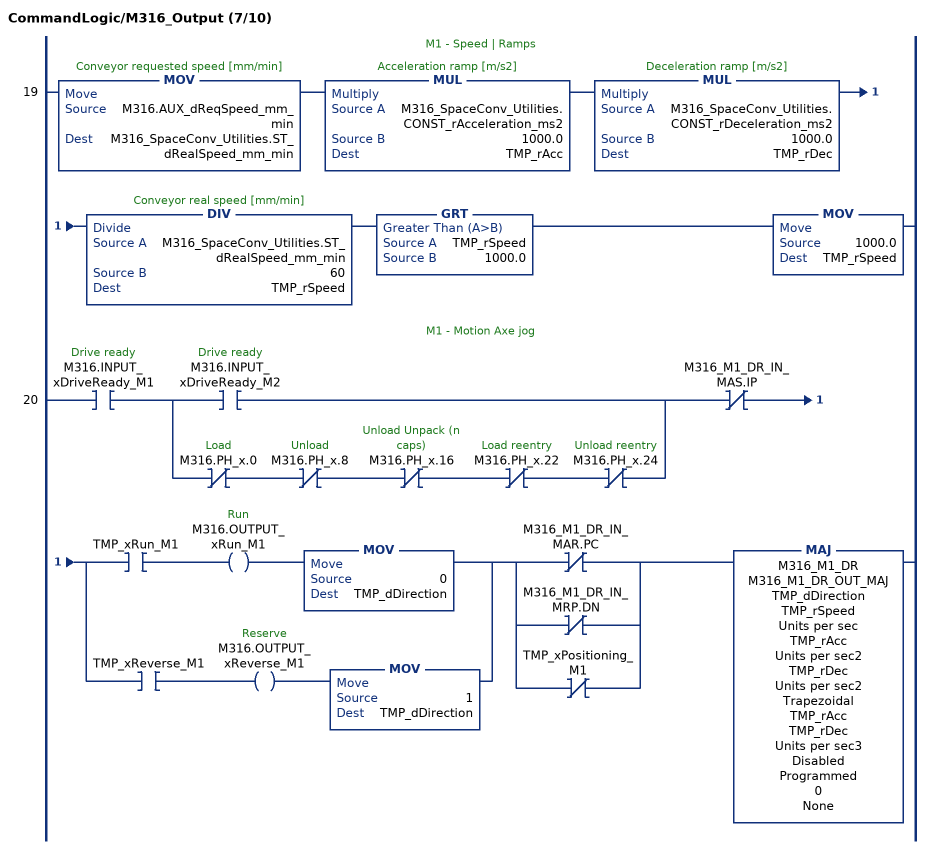
   // M1 - Speed | Ramps
   19: MOV(M316.AUX_dReqSpeed_mm_min,M316_SpaceConv_Utilities.ST_dRealSpeed_mm_min)MUL(M316_SpaceConv_Utilities.CONST_rAcceleration_ms2,1000.0,TMP_rAcc)MUL(M316_SpaceConv_Utilities.CONST_rDeceleration_ms2,1000.0,TMP_rDec)DIV(M316_SpaceConv_Utilities.ST_dRealSpeed_mm_min,60,TMP_rSpeed)GRT(TMP_rSpeed,1000.0)MOV(1000.0,TMP_rSpeed);
   // M1 - Motion Axe jog
   20: XIC(M316.INPUT_xDriveReady_M1)[XIC(M316.INPUT_xDriveReady_M2) ,XIO(M316.PH_x.0) XIO(M316.PH_x.8) XIO(M316.PH_x.16) XIO(M316.PH_x.22) XIO(M316.PH_x.24) ]XIO(M316_M1_DR_IN_MAS.IP)[XIC(TMP_xRun_M1) OTE(M316.OUTPUT_xRun_M1) MOV(0,TMP_dDirection) ,XIC(TMP_xReverse_M1) OTE(M316.OUTPUT_xReverse_M1) MOV(1,TMP_dDirection) ][XIO(M316_M1_DR_IN_MAR.PC) ,XIO(M316_M1_DR_IN_MRP.DN) ,XIO(TMP_xPositioning_M1) ]MAJ(M316_M1_DR,M316_M1_DR_OUT_MAJ,TMP_dDirection,TMP_rSpeed,Units per sec,TMP_rAcc,Units per sec2,TMP_rDec,Units per sec2,Trapezoidal,TMP_rAcc,TMP_rDec,Units per sec3,Disabled,Programmed,0,None);
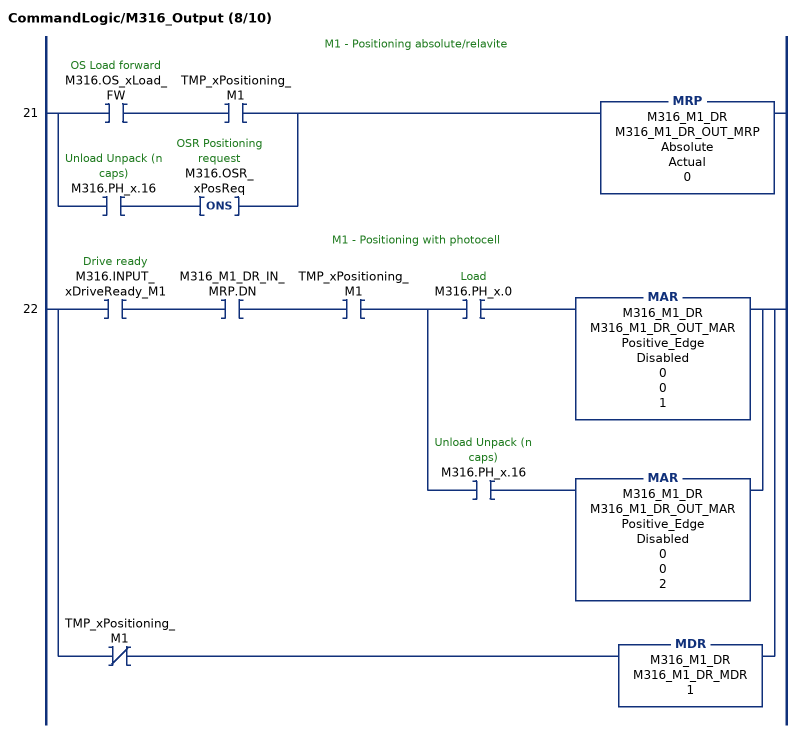
   // M1 - Positioning absolute/relavite
   21: [XIC(M316.OS_xLoad_FW) XIC(TMP_xPositioning_M1) ,XIC(M316.PH_x.16) ONS(M316.OSR_xPosReq) ]MRP(M316_M1_DR,M316_M1_DR_OUT_MRP,Absolute,Actual,0);
   // M1 - Positioning with photocell
   22: [XIC(M316.INPUT_xDriveReady_M1) XIC(M316_M1_DR_IN_MRP.DN) XIC(TMP_xPositioning_M1) [XIC(M316.PH_x.0) MAR(M316_M1_DR,M316_M1_DR_OUT_MAR,Positive_Edge,Disabled,0,0,1) ,XIC(M316.PH_x.16) MAR(M316_M1_DR,M316_M1_DR_OUT_MAR,Positive_Edge,Disabled,0,0,2) ] ,XIO(TMP_xPositioning_M1) MDR(M316_M1_DR,M316_M1_DR_MDR,1) ];
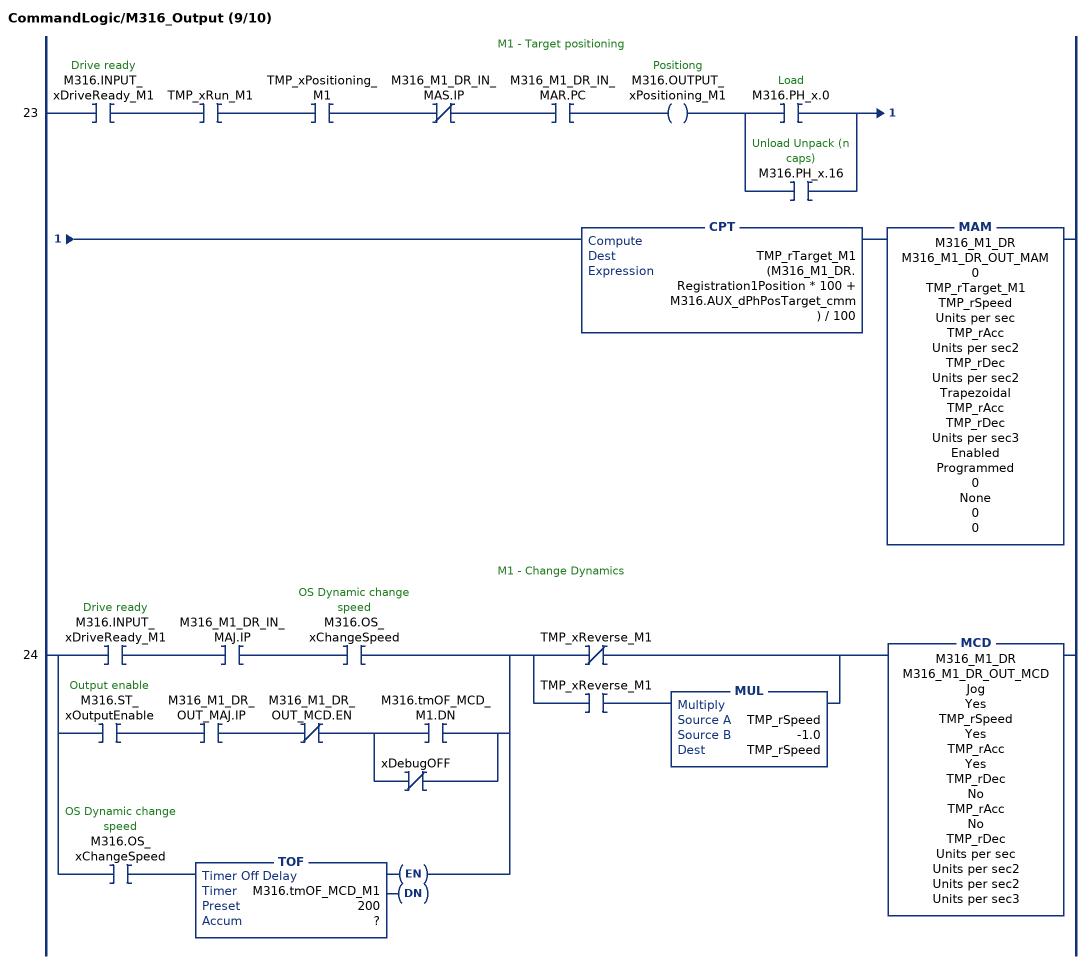
   // M1 - Target positioning
   23: XIC(M316.INPUT_xDriveReady_M1)XIC(TMP_xRun_M1)XIC(TMP_xPositioning_M1)XIO(M316_M1_DR_IN_MAS.IP)XIC(M316_M1_DR_IN_MAR.PC)OTE(M316.OUTPUT_xPositioning_M1)[XIC(M316.PH_x.0) ,XIC(M316.PH_x.16) ]CPT(TMP_rTarget_M1,(M316_M1_DR.Registration1Position * 100 + M316.AUX_dPhPosTarget_cmm ) / 100)MAM(M316_M1_DR,M316_M1_DR_OUT_MAM,0,TMP_rTarget_M1,TMP_rSpeed,Units per sec,TMP_rAcc,Units per sec2,TMP_rDec,Units per sec2,Trapezoidal,TMP_rAcc,TMP_rDec,Units per sec3,Enabled,Programmed,0,None,0,0);
   // M1 - Change Dynamics
   24: [XIC(M316.INPUT_xDriveReady_M1) XIC(M316_M1_DR_IN_MAJ.IP) XIC(M316.OS_xChangeSpeed) ,XIC(M316.ST_xOutputEnable) XIC(M316_M1_DR_OUT_MAJ.IP) XIO(M316_M1_DR_OUT_MCD.EN) [XIC(M316.tmOF_MCD_M1.DN) ,XIO(xDebugOFF) ] ,XIC(M316.OS_xChangeSpeed) TOF(M316.tmOF_MCD_M1,?,?) ][XIO(TMP_xReverse_M1) ,XIC(TMP_xReverse_M1) MUL(TMP_rSpeed,-1.0,TMP_rSpeed) ]MCD(M316_M1_DR,M316_M1_DR_OUT_MCD,Jog,Yes,TMP_rSpeed,Yes,TMP_rAcc,Yes,TMP_rDec,No,TMP_rAcc,No,TMP_rDec,Units per sec,Units per sec2,Units per sec2,Units per sec3);
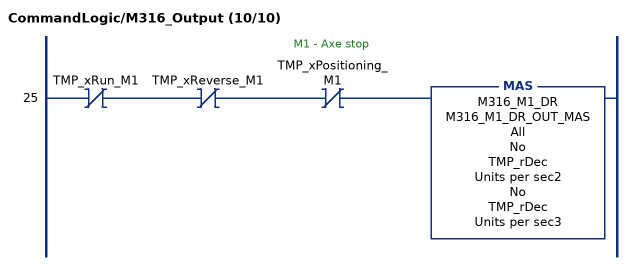
   // M1 - Axe stop
   25: XIO(TMP_xRun_M1)XIO(TMP_xReverse_M1)XIO(TMP_xPositioning_M1)MAS(M316_M1_DR,M316_M1_DR_OUT_MAS,All,No,TMP_rDec,Units per sec2,No,TMP_rDec,Units per sec3);
END_ROUTINE

ROUTINE M316A_Output   (* ladder *)
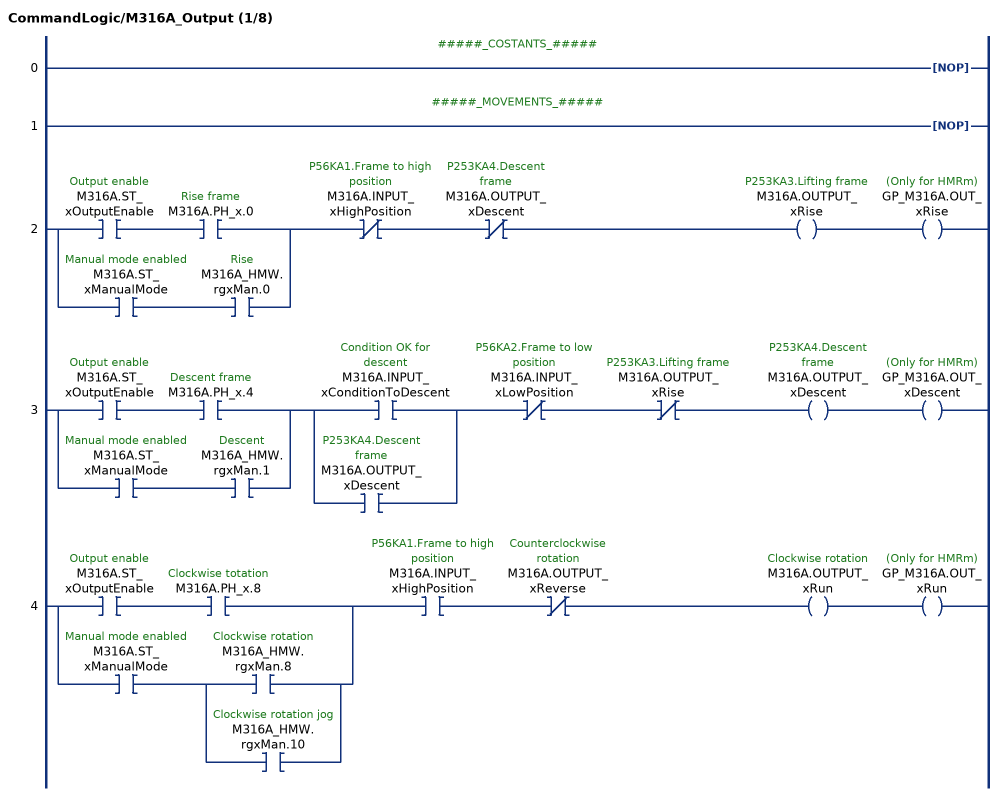
   // #####_COSTANTS_#####
   0: NOP();
   // #####_MOVEMENTS_#####
   1: NOP();
   2: [XIC(M316A.ST_xOutputEnable) XIC(M316A.PH_x.0) ,XIC(M316A.ST_xManualMode) XIC(M316A_HMW.rgxMan.0) ]XIO(M316A.INPUT_xHighPosition)XIO(M316A.OUTPUT_xDescent)OTE(M316A.OUTPUT_xRise)OTE(GP_M316A.OUT_xRise);
   3: [XIC(M316A.ST_xOutputEnable) XIC(M316A.PH_x.4) ,XIC(M316A.ST_xManualMode) XIC(M316A_HMW.rgxMan.1) ][XIC(M316A.INPUT_xConditionToDescent) ,XIC(M316A.OUTPUT_xDescent) ]XIO(M316A.INPUT_xLowPosition)XIO(M316A.OUTPUT_xRise)OTE(M316A.OUTPUT_xDescent)OTE(GP_M316A.OUT_xDescent);
   4: [XIC(M316A.ST_xOutputEnable) XIC(M316A.PH_x.8) ,XIC(M316A.ST_xManualMode) [XIC(M316A_HMW.rgxMan.8) ,XIC(M316A_HMW.rgxMan.10) ] ]XIC(M316A.INPUT_xHighPosition)XIO(M316A.OUTPUT_xReverse)OTE(M316A.OUTPUT_xRun)OTE(GP_M316A.OUT_xRun);
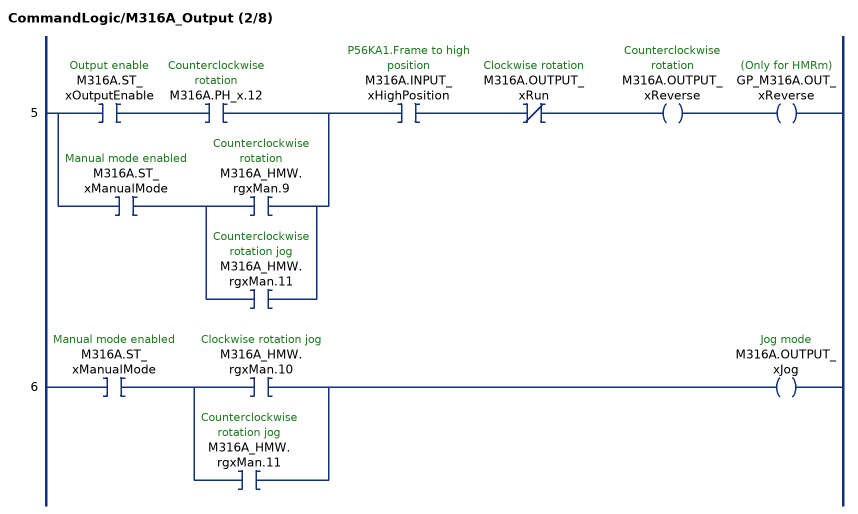
   5: [XIC(M316A.ST_xOutputEnable) XIC(M316A.PH_x.12) ,XIC(M316A.ST_xManualMode) [XIC(M316A_HMW.rgxMan.9) ,XIC(M316A_HMW.rgxMan.11) ] ]XIC(M316A.INPUT_xHighPosition)XIO(M316A.OUTPUT_xRun)OTE(M316A.OUTPUT_xReverse)OTE(GP_M316A.OUT_xReverse);
   6: XIC(M316A.ST_xManualMode)[XIC(M316A_HMW.rgxMan.10) ,XIC(M316A_HMW.rgxMan.11) ]OTE(M316A.OUTPUT_xJog);
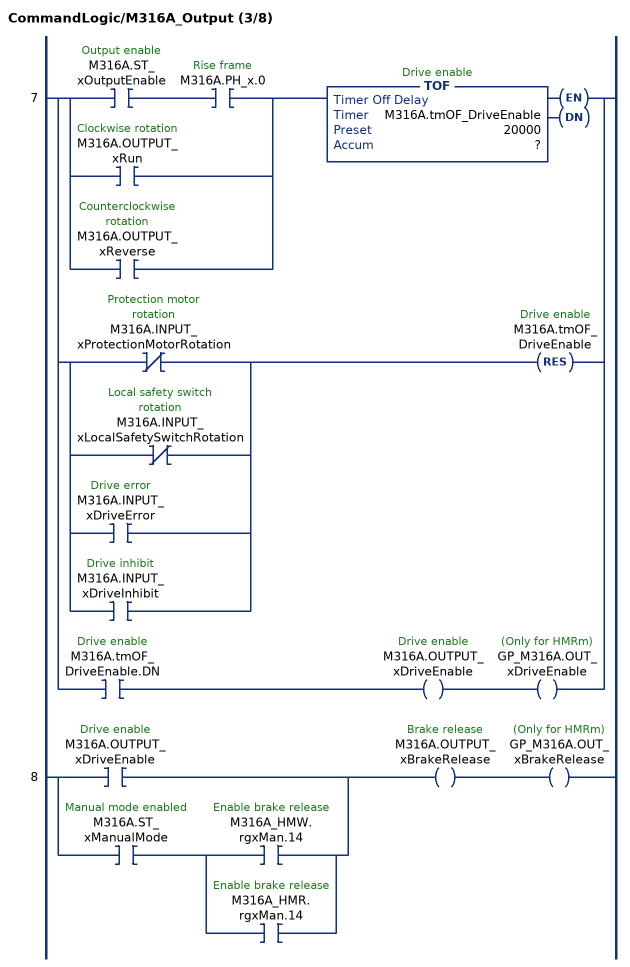
   7: [[XIC(M316A.ST_xOutputEnable) XIC(M316A.PH_x.0) ,XIC(M316A.OUTPUT_xRun) ,XIC(M316A.OUTPUT_xReverse) ] TOF(M316A.tmOF_DriveEnable,?,?) ,[XIO(M316A.INPUT_xProtectionMotorRotation) ,XIO(M316A.INPUT_xLocalSafetySwitchRotation) ,XIC(M316A.INPUT_xDriveError) ,XIC(M316A.INPUT_xDriveInhibit) ] RES(M316A.tmOF_DriveEnable) ,XIC(M316A.tmOF_DriveEnable.DN) OTE(M316A.OUTPUT_xDriveEnable) OTE(GP_M316A.OUT_xDriveEnable) ];
   8: [XIC(M316A.OUTPUT_xDriveEnable) ,XIC(M316A.ST_xManualMode) [XIC(M316A_HMW.rgxMan.14) ,XIC(M316A_HMR.rgxMan.14) ] ]OTE(M316A.OUTPUT_xBrakeRelease)OTE(GP_M316A.OUT_xBrakeRelease);
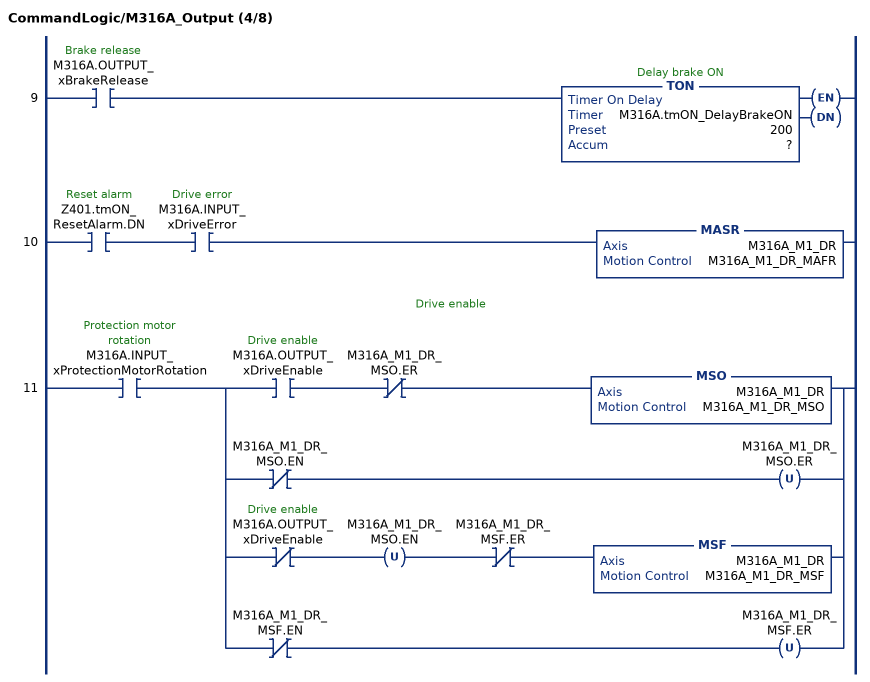
   9: XIC(M316A.OUTPUT_xBrakeRelease)TON(M316A.tmON_DelayBrakeON,?,?);
   10: XIC(Z401.tmON_ResetAlarm.DN)XIC(M316A.INPUT_xDriveError)MASR(M316A_M1_DR,M316A_M1_DR_MAFR);
   // Drive enable
   11: XIC(M316A.INPUT_xProtectionMotorRotation)[XIC(M316A.OUTPUT_xDriveEnable) XIO(M316A_M1_DR_MSO.ER) MSO(M316A_M1_DR,M316A_M1_DR_MSO) ,XIO(M316A_M1_DR_MSO.EN) OTU(M316A_M1_DR_MSO.ER) ,XIO(M316A.OUTPUT_xDriveEnable) OTU(M316A_M1_DR_MSO.EN) XIO(M316A_M1_DR_MSF.ER) MSF(M316A_M1_DR,M316A_M1_DR_MSF) ,XIO(M316A_M1_DR_MSF.EN) OTU(M316A_M1_DR_MSF.ER) ];
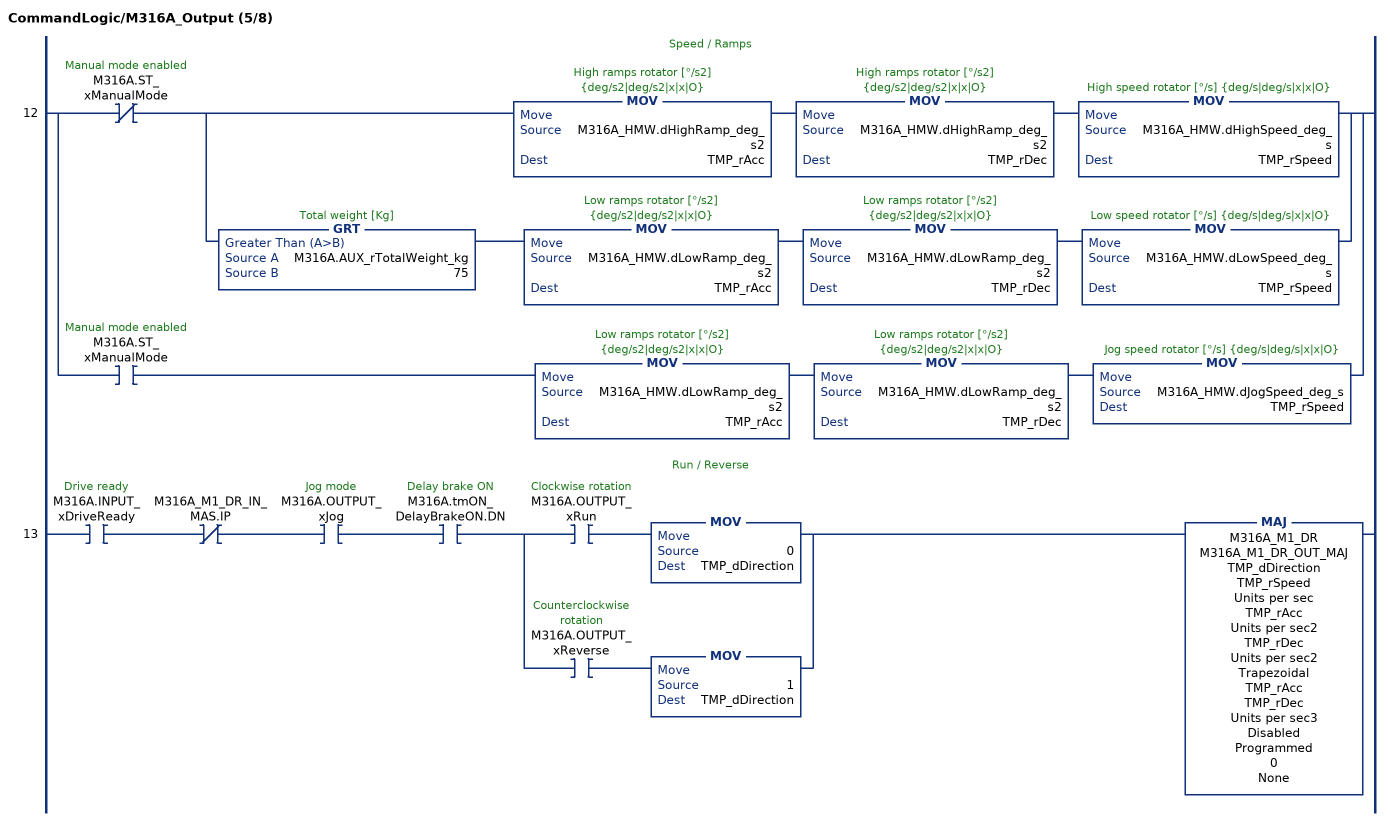
   // Speed / Ramps
   12: [XIO(M316A.ST_xManualMode) [MOV(M316A_HMW.dHighRamp_deg_s2,TMP_rAcc) MOV(M316A_HMW.dHighRamp_deg_s2,TMP_rDec) MOV(M316A_HMW.dHighSpeed_deg_s,TMP_rSpeed) ,GRT(M316A.AUX_rTotalWeight_kg,75) MOV(M316A_HMW.dLowRamp_deg_s2,TMP_rAcc) MOV(M316A_HMW.dLowRamp_deg_s2,TMP_rDec) MOV(M316A_HMW.dLowSpeed_deg_s,TMP_rSpeed) ] ,XIC(M316A.ST_xManualMode) MOV(M316A_HMW.dLowRamp_deg_s2,TMP_rAcc) MOV(M316A_HMW.dLowRamp_deg_s2,TMP_rDec) MOV(M316A_HMW.dJogSpeed_deg_s,TMP_rSpeed) ];
   // Run / Reverse
   13: XIC(M316A.INPUT_xDriveReady)XIO(M316A_M1_DR_IN_MAS.IP)XIC(M316A.OUTPUT_xJog)XIC(M316A.tmON_DelayBrakeON.DN)[XIC(M316A.OUTPUT_xRun) MOV(0,TMP_dDirection) ,XIC(M316A.OUTPUT_xReverse) MOV(1,TMP_dDirection) ]MAJ(M316A_M1_DR,M316A_M1_DR_OUT_MAJ,TMP_dDirection,TMP_rSpeed,Units per sec,TMP_rAcc,Units per sec2,TMP_rDec,Units per sec2,Trapezoidal,TMP_rAcc,TMP_rDec,Units per sec3,Disabled,Programmed,0,None);
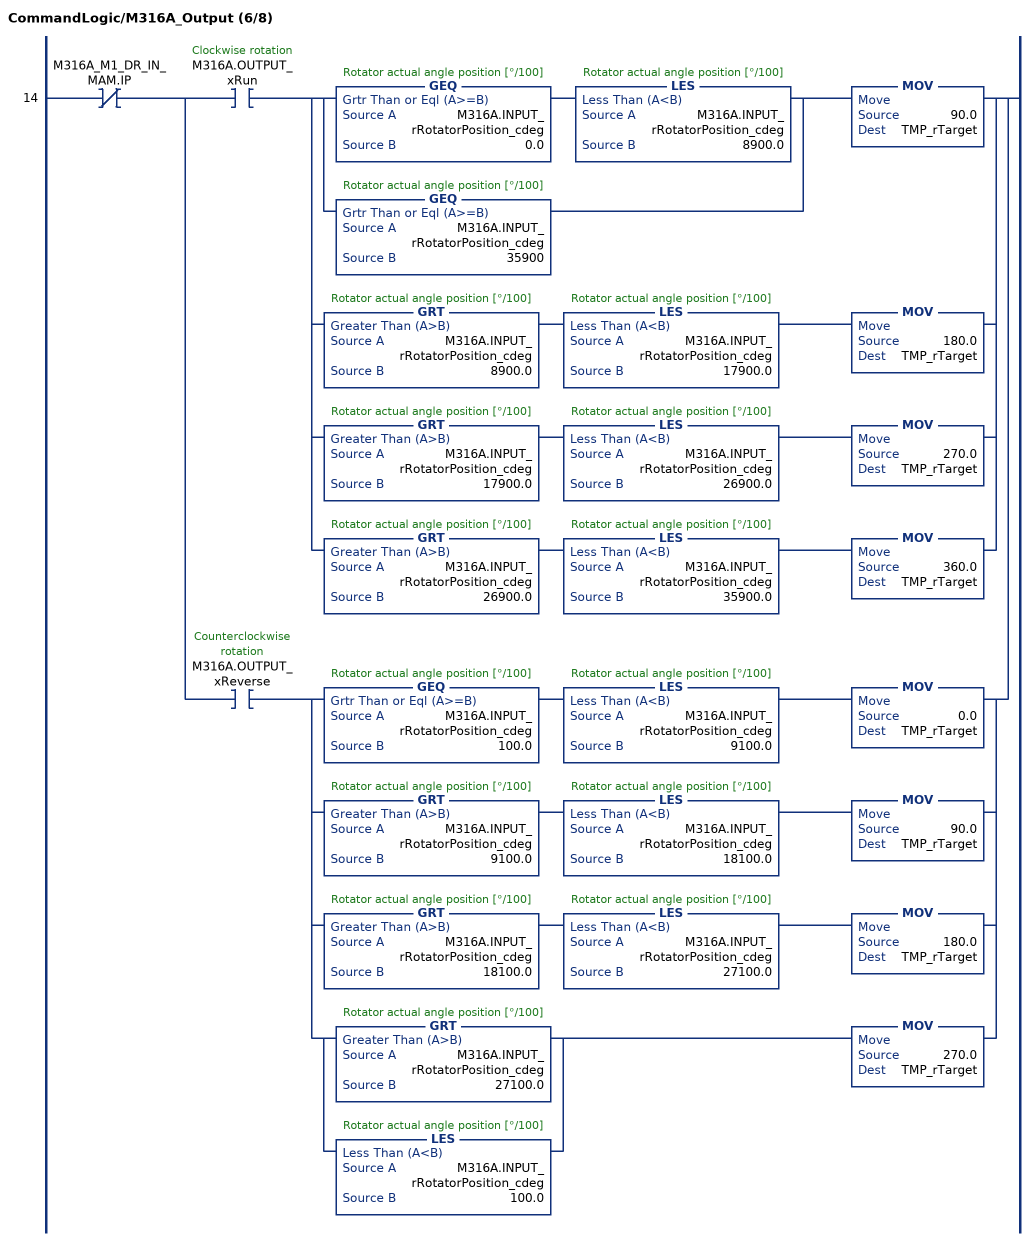
   14: XIO(M316A_M1_DR_IN_MAM.IP)[XIC(M316A.OUTPUT_xRun) [[GEQ(M316A.INPUT_rRotatorPosition_cdeg,0.0) LES(M316A.INPUT_rRotatorPosition_cdeg,8900.0) ,GEQ(M316A.INPUT_rRotatorPosition_cdeg,35900) ] MOV(90.0,TMP_rTarget) ,GRT(M316A.INPUT_rRotatorPosition_cdeg,8900.0) LES(M316A.INPUT_rRotatorPosition_cdeg,17900.0) MOV(180.0,TMP_rTarget) ,GRT(M316A.INPUT_rRotatorPosition_cdeg,17900.0) LES(M316A.INPUT_rRotatorPosition_cdeg,26900.0) MOV(270.0,TMP_rTarget) ,GRT(M316A.INPUT_rRotatorPosition_cdeg,26900.0) LES(M316A.INPUT_rRotatorPosition_cdeg,35900.0) MOV(360.0,TMP_rTarget) ] ,XIC(M316A.OUTPUT_xReverse) [GEQ(M316A.INPUT_rRotatorPosition_cdeg,100.0) LES(M316A.INPUT_rRotatorPosition_cdeg,9100.0) MOV(0.0,TMP_rTarget) ,GRT(M316A.INPUT_rRotatorPosition_cdeg,9100.0) LES(M316A.INPUT_rRotatorPosition_cdeg,18100.0) MOV(90.0,TMP_rTarget) ,GRT(M316A.INPUT_rRotatorPosition_cdeg,18100.0) LES(M316A.INPUT_rRotatorPosition_cdeg,27100.0) MOV(180.0,TMP_rTarget) ,[GRT(M316A.INPUT_rRotatorPosition_cdeg,27100.0) ,LES(M316A.INPUT_rRotatorPosition_cdeg,100.0) ] MOV(270.0,TMP_rTarget) ] ];
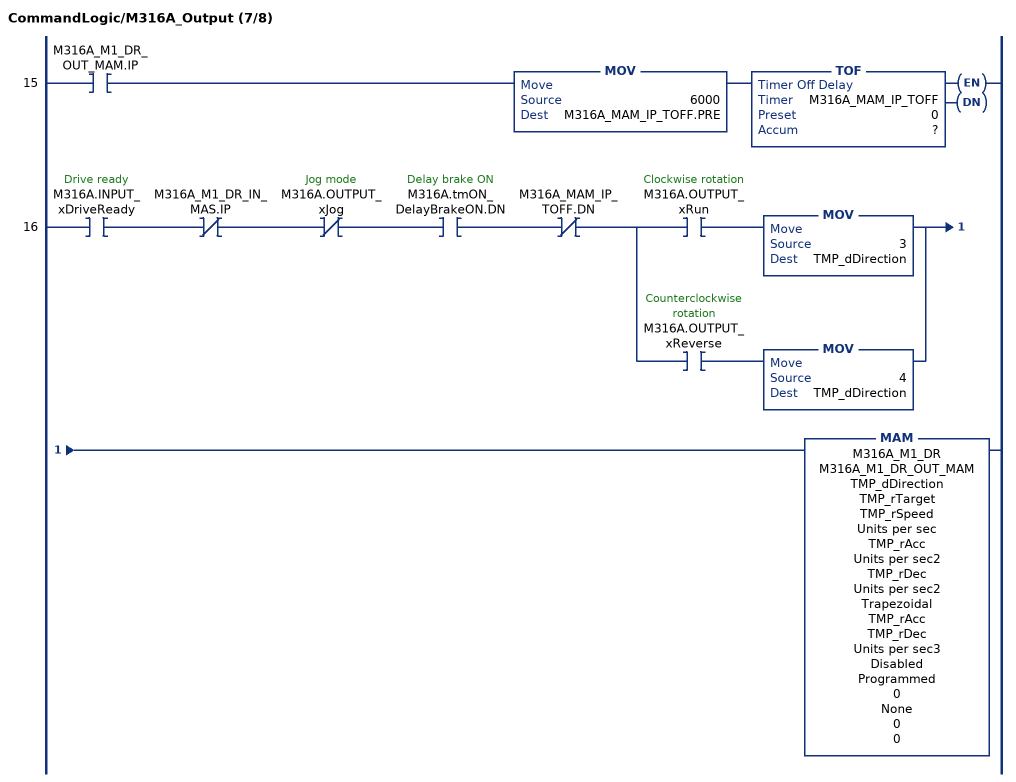
   15: XIC(M316A_M1_DR_OUT_MAM.IP)MOV(6000,M316A_MAM_IP_TOFF.PRE)TOF(M316A_MAM_IP_TOFF,?,?);
   16: XIC(M316A.INPUT_xDriveReady)XIO(M316A_M1_DR_IN_MAS.IP)XIO(M316A.OUTPUT_xJog)XIC(M316A.tmON_DelayBrakeON.DN)XIO(M316A_MAM_IP_TOFF.DN)[XIC(M316A.OUTPUT_xRun) MOV(3,TMP_dDirection) ,XIC(M316A.OUTPUT_xReverse) MOV(4,TMP_dDirection) ]MAM(M316A_M1_DR,M316A_M1_DR_OUT_MAM,TMP_dDirection,TMP_rTarget,TMP_rSpeed,Units per sec,TMP_rAcc,Units per sec2,TMP_rDec,Units per sec2,Trapezoidal,TMP_rAcc,TMP_rDec,Units per sec3,Disabled,Programmed,0,None,0,0);
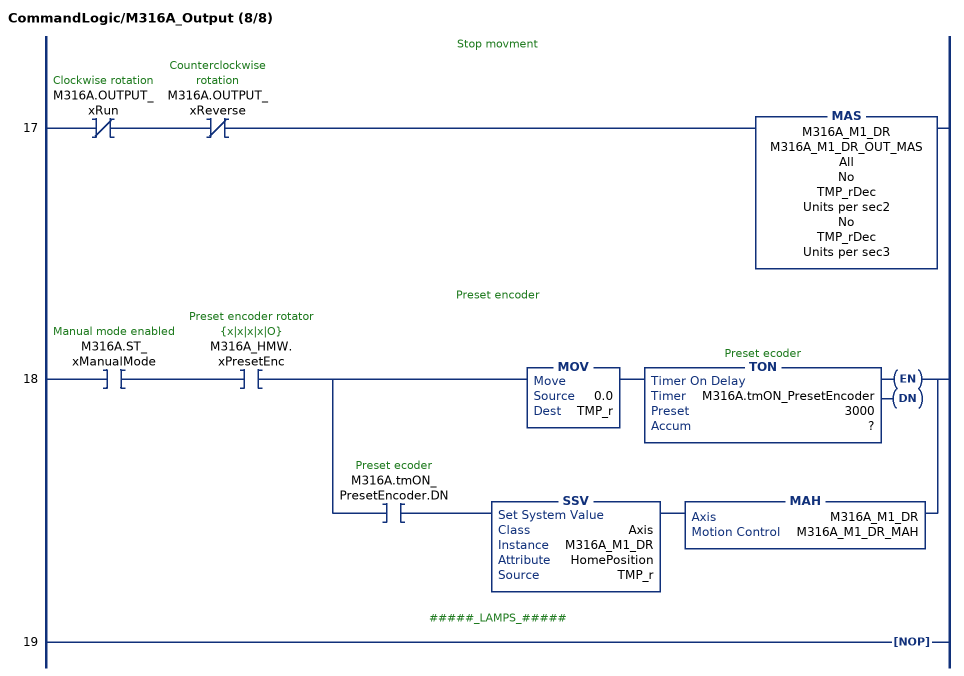
   // Stop movment
   17: XIO(M316A.OUTPUT_xRun)XIO(M316A.OUTPUT_xReverse)MAS(M316A_M1_DR,M316A_M1_DR_OUT_MAS,All,No,TMP_rDec,Units per sec2,No,TMP_rDec,Units per sec3);
   // Preset encoder
   18: XIC(M316A.ST_xManualMode)XIC(M316A_HMW.xPresetEnc)[MOV(0.0,TMP_r) TON(M316A.tmON_PresetEncoder,?,?) ,XIC(M316A.tmON_PresetEncoder.DN) SSV(Axis,M316A_M1_DR,HomePosition,TMP_r) MAH(M316A_M1_DR,M316A_M1_DR_MAH) ];
   // #####_LAMPS_#####
   19: NOP();
END_ROUTINE
